REGION Network 3: Release drive
   //
         O     #Temp_IO_Status.Switch_Drive_ON_OFF;
         O     #IN_Request_Filling;
         O     #IN_Request_Feedpump;
         O     #IN_Request_Cooling;
         O     #IN_Request_Heating;
         A     #IN_Release;
         =     #Temp_ReleaseDrive;
END_REGION

REGION Network 4: Faults
         A     #IN_Reset_fault;
         R     #Temp_IO_Fault.FLT_Motorprotection;
         R     #Temp_IO_Fault.FLT_FrequencyConverter;
         R     #Temp_IO_Fault.FLT_MaxP_MaxLTripTray;
         R     #Temp_IO_Fault.FLT_Dryrunsafety;
         R     #Temp_IO_Fault.FLT_wrong_Timevalue;

         A     #IN_Fault_Motorprotection;
         S     #Temp_IO_Fault.FLT_Motorprotection;
         S     #Temp_IO_Status.Reset_Intervall;
   //
         A     #IN_ControlVoltage;
         AN    #Temp_IO_Fault.FLT_wrong_Timevalue;
         AN    #Temp_IO_Status.Start_Startupdelay;
         L     S5T#5S;
         SD    #IN_TimerStartUpFConv;
   //
         A     #IN_TimerStartUpFConv;
         AN    #IN_FaultFreqConverter;
         A     #Temp_ReleaseDrive;
         A     #Temp_IO_Status.Config_bit_with_FC;
         S     #Temp_IO_Fault.FLT_FrequencyConverter;
         S     #Temp_IO_Status.Reset_Intervall;
   //
         AN    #IN_MaxPressure_MaxLTray;
         A     #Temp_ReleaseDrive;
         S     #Temp_IO_Fault.FLT_MaxP_MaxLTripTray;
         S     #Temp_IO_Status.Reset_Intervall;
   //
         AN    #IN_DryRun;
         A     #Temp_ReleaseDrive;
         S     #Temp_IO_Fault.FLT_Dryrunsafety;
         S     #Temp_IO_Status.Reset_Intervall;
END_REGION

REGION Network 5: Time handle
   // Es werden die Absolutwerte der Zeiten berechnet um sie dann vergleichen zu 
   // können. Intervallzeiten sind minimal 10sec. Sonst Störung "Zeitwert falsch"!
   // Bei Spaltfiltern max Laufzeit 20sec.,Min Pausenzeit 300sec.und kein Dauerbetrieb
   // möglich!
         SET;
         R     #Temp_IO_Fault.FLT_wrong_Timevalue;
   //
         L     #IN_DW_RunTime;
         T     #Temp_RunTime;
         L     #IN_DW_PauseTime;
         T     #Temp_PauseTime;
   //
   // Absolutwerte berechnen
   //
         CALL  T_CONV
         ( IN  := #Temp_RunTime,
           OUT := #Temp_Runtime_ms
         );
   //
         CALL  T_CONV
         ( IN  := #Temp_PauseTime,
           OUT := #Temp_Pausetime_ms
         );
   //
         SET;
         R     #Temp_IO_Status.No_Pausetime;
   //
         L     #Temp_Runtime_ms;
         L     0;
         ==I;
         O(;
         L     #Temp_Pausetime_ms;
         L     0;
         ==I;
         );
         AN    #Temp_IO_Status.Config_bit_split;  // Bei Spaltfilter immer mit Intervall
         S     #Temp_IO_Status.No_Pausetime;
   //
   // Zeiten limitieren
   //
         A     #Temp_IO_Status.Config_bit_split;  // Bei Spaltfilter Kontrolle auf spezielle Min und Maxwerte
         JC    nLi2;
   //
         L     #Temp_Runtime_ms;
         L     10000;  // 10 sec
         <D;
         S     #Temp_IO_Fault.FLT_wrong_Timevalue;  // Antrieb STOP!!!
         JCN   nLi1;
         L     S5T#10S;
         T     #Temp_RunTime;
   //
   nLi1: L     #Temp_Pausetime_ms;
         L     10000;  // 10.0 sec
         <D;
         S     #Temp_IO_Fault.FLT_wrong_Timevalue;  // Antrieb STOP!!!
         JCN   nLi3;
         L     S5T#10S;
         T     #Temp_PauseTime;
         JU    nLi3;
   //
   // Sonderteil für Spaltfilter
   nLi2: L     #Temp_Runtime_ms;
         L     20000;  // 20.0 sec
         >D;
         S     #Temp_IO_Fault.FLT_wrong_Timevalue;  // Antrieb STOP!!!
         JCN   KfS1;
         L     S5T#20S;
         T     #Temp_RunTime;
   KfS1: L     #Temp_Pausetime_ms;
         L     L#300000;  // 300.0 sec
         <D;
         S     #Temp_IO_Fault.FLT_wrong_Timevalue;  // Antrieb STOP!!!
         JCN   nLi3;
         L     S5T#5M;
         T     #Temp_PauseTime;
   //
   nLi3: NOP   0;
         A     #Temp_IO_Status.No_Pausetime;  // Wenn eh eine zeit null dann andere egal!
         R     #Temp_IO_Fault.FLT_wrong_Timevalue;
END_REGION

REGION Network 6: Reset Intervall / Angefordert setzen
         O     #Temp_IO_Status.No_Pausetime;
         S     #Temp_IO_Status.Reset_Intervall;
   //
         ON    #Temp_ReleaseDrive;
         ON    #IN_Release;
         O     #Temp_IO_Status.Reset_Intervall;
         R     #Temp_IO_Status.Run;
         R     #Temp_IO_Status.Pause;
         R     #Temp_IO_Status.Reset_Intervall;
END_REGION

REGION Network 7: Wiedereinschaltsperre
         ON    #IN_ControlVoltage;
         FP    #Temp_IO_Status.Ramp_CVoltage_Off;
         S     #Temp_IO_Status.Start_Startupdelay;
         R     #Temp_IO_Status.Disable_Start;
         R     #IN_TimerDrive;
   //
         ON    #Temp_IO_Status.Config_bit_with_FC;
         O     #IN_TimerDrive;
         A     #Temp_IO_Status.Start_Startupdelay;
         R     #Temp_IO_Status.Disable_Start;
         R     #Temp_IO_Status.Start_Startupdelay;
   //
         A     #Temp_IO_Status.Start_Startupdelay;
         JCN   Lauf;
   //
         A     #Temp_IO_Status.Disable_Start;
         L     S5T#10S;
         SD    #IN_TimerDrive;
   //
         SET;
         S     #Temp_IO_Status.Disable_Start;
   //
         A     #IN_TimerDrive;
         A     #Temp_IO_Status.Start_Startupdelay;
         R     #Temp_IO_Status.Start_Startupdelay;
         R     #Temp_IO_Status.Disable_Start;
END_REGION

REGION Network 8: Laufzeit
   Lauf: NOP   0;
         A     #Temp_ReleaseDrive;
         AN    #Temp_IO_Status.Pause;
         AN    #Temp_IO_Status.Start_Startupdelay;
         JCN   Paus;
   //
         A     #Temp_IO_Status.Run;
         L     #Temp_RunTime;
         SD    #IN_TimerDrive;
   //
         SET;
         S     #Temp_IO_Status.Run;
   //
         A     #IN_TimerDrive;
         JCN   Ausg;
         SET;
         R     #Temp_IO_Status.Run;
         R     #IN_TimerDrive;
END_REGION

REGION Network 9: Pause
   Paus: NOP   0;
         A     #Temp_ReleaseDrive;
         AN    #Temp_IO_Status.Run;
         AN    #Temp_IO_Status.Start_Startupdelay;
         JCN   Ausg;
   //
         A     #Temp_IO_Status.Pause;
         L     #Temp_PauseTime;
         SD    #IN_TimerDrive;
   //
         SET;
         S     #Temp_IO_Status.Pause;
   //
         A     #IN_TimerDrive;
         JCN   Ausg;
         SET;
         R     #Temp_IO_Status.Pause;
         R     #IN_TimerDrive;
END_REGION

REGION Network 10: Output mainscontactor
   Ausg: NOP   0;
   //
         A(;
   //
         A     #IN_ControlVoltage;  // generell Eingeschaltet mit FU
         A     #Temp_IO_Status.Config_bit_with_FC;
         AN    #Temp_IO_Status.Start_Startupdelay;
   //
         O(;
         A     #Temp_IO_Status.Run;  // generell Eingeschaltet ohne FU
         O     #Temp_IO_Status.No_Pausetime;
         A     #Temp_IO_Status.Switch_Drive_ON_OFF;
         A(;
         AN    #Temp_IO_Fault.FLT_Dryrunsafety;
         O     #Temp_IO_Status.Config_bit_split;
         );
         AN    #Temp_IO_Status.Config_bit_with_FC;
         );
   //
         O(;
         A     #IN_Request_Filling;  // Befuellen als Füllpumpe
         A     #Temp_IO_Status.Config_bit_char;
         );
   //
         O(;
         O     #Temp_IO_Status.No_Pausetime;  // Befuellen aber normal konfiguriert
         O     #Temp_IO_Status.Run;
         A     #IN_Request_Filling;
         AN    #Temp_IO_Fault.FLT_Dryrunsafety;
         A     #Temp_IO_Status.Config_bit_normal;
         );
   //
         O(;
         A     #IN_Request_Filling;  // aber auch beim Befüllen
         AN    #Temp_IO_Fault.FLT_Dryrunsafety;
         A     #Temp_IO_Status.Run;
         O     #IN_Request_Feedpump;  // Speisen
         A     #Temp_IO_Status.config_bit_feed;
         );
   //
         O(;
         A     #IN_Request_Heating;  // Beim Heizen mit Intervall
         A(;
         O     #Temp_IO_Status.Run;
         O     #Temp_IO_Status.No_Pausetime;
         );
         O     #IN_Request_Cooling;  // Kühlen ohne Intervall, damit WT nicht einfriert
         AN    #Temp_IO_Status.Config_bit_with_FC;
         AN    #Temp_IO_Status.Config_bit_split;
         AN    #Temp_IO_Fault.FLT_Dryrunsafety;
         );
   //
         );
   //
         A(;
         A     #IN_Release;
         AN    #Temp_IO_Fault.FLT_wrong_Timevalue;
         AN    #Temp_IO_Fault.FLT_MaxP_MaxLTripTray;
         O     #Temp_IO_Status.Config_bit_with_FC;  // Wenn FU dann immer an!
         );
         AN    #Temp_IO_Fault.FLT_Motorprotection;
         AN    #Temp_IO_Fault.FLT_Dryrunsafety;
   //
         =     #OUT_MainsContactor;
         =     #Temp_MainsContactor;
END_REGION

REGION Network 11: Ouput release frequency converter
         O     #Temp_IO_Status.No_Pausetime;
         O     #Temp_IO_Status.Run;
         O     #IN_Request_Feedpump;
         A     #IN_Release;
         A     #Temp_MainsContactor;
         A     #Temp_IO_Status.Config_bit_with_FC;
         A(;
         O     #Temp_IO_Status.Switch_Drive_ON_OFF;
         O     #IN_Request_Feedpump;
         );
         AN    #Temp_IO_Fault.FLT_FrequencyConverter;
         A     #IN_FaultFreqConverter;
         =     #OUT_Release_FConverter;
         =     #Temp_Release_FConverter;
END_REGION

REGION Network 12: Error handling
         O     #Temp_IO_Fault.FLT_Motorprotection;
         O     #Temp_IO_Fault.FLT_FrequencyConverter;
         O     #Temp_IO_Fault.FLT_MaxP_MaxLTripTray;
         O     #Temp_IO_Fault.FLT_Dryrunsafety;
         O     #Temp_IO_Fault.FLT_wrong_Timevalue;
         =     #Temp_Fault_Drive;
         =     #Temp_IO_Status.FaultExist;

         O     #Temp_IO_Fault.FLT_Motorprotection;
         O     #Temp_IO_Fault.FLT_FrequencyConverter;
         O     #Temp_IO_Fault.FLT_Dryrunsafety;
         A     #IN_SelectFaultLevel;
         S     #IO_FaultLevel_1;

         O     #Temp_IO_Fault.FLT_Motorprotection;
         O     #Temp_IO_Fault.FLT_FrequencyConverter;
         O     #Temp_IO_Fault.FLT_Dryrunsafety;
         AN    #IN_SelectFaultLevel;
         O;
         O     #Temp_IO_Fault.FLT_MaxP_MaxLTripTray;
         O     #Temp_IO_Fault.FLT_wrong_Timevalue;
         S     #IO_FaultLevel_3;

         O     #Temp_IO_Fault.FLT_Motorprotection;
         FP    #Temp_IO_Status.FLT_Motorprotection;
         S     #IO_NewFault;

         O     #Temp_IO_Fault.FLT_FrequencyConverter;
         FP    #Temp_IO_Status.FLT_FC;
         S     #IO_NewFault;

         O     #Temp_IO_Fault.FLT_MaxP_MaxLTripTray;
         FP    #Temp_IO_Status.FLT_MaxP_MaxLTripTray;
         S     #IO_NewFault;

         O     #Temp_IO_Fault.FLT_Dryrunsafety;
         FP    #Temp_IO_Status.FLT_Dryrunsafety;
         S     #IO_NewFault;

         O     #Temp_IO_Fault.FLT_wrong_Timevalue;
         FP    #Temp_IO_Status.FLT_wrong_Timevalue;
         S     #IO_NewFault;
END_REGION

REGION Network 13: State of drive: 1-> ON; 2->Faulty; 3->Selected but not on
         L     0;
         O     #Temp_Fault_Drive;
         JCN   err;
         L     2;
         JU    tran;
   err:  AN    #Temp_IO_Status.Config_bit_with_FC;
         A     #Temp_MainsContactor;
         O     #Temp_Release_FConverter;
         JCN   anl;
         L     1;
         JU    tran;
   anl:  AN    #Temp_IO_Status.Config_bit_with_FC;
         A     #Temp_MainsContactor;
         O     #Temp_Release_FConverter;
         ON    #Temp_IO_Status.Switch_Drive_ON_OFF;
         JC    tran;
         L     3;
   tran: T     #Temp_IO_Status.State_Drive;
END_REGION

REGION Network 14: Save data
         CALL  BLKMOV
         ( SRCBLK  := #Temp_IO_Status,
           RET_VAL := #ERROR_CODE,
           DSTBLK  := #Anyzeiger1
         );
   //
         CALL  BLKMOV
         ( SRCBLK  := #Temp_IO_Fault,
           RET_VAL := #ERROR_CODE,
           DSTBLK  := #Anyzeiger2
         );
   //
END_REGION
END_FUNCTION

FUNCTION "FC102_Refilling" : Void   // FC102, STL
TITLE = Filling of a tank
{ S7_Optimized_Access := 'FALSE' }
AUTHOR : KT242
FAMILY : RS_KK
NAME : Filling
VERSION : 1.1
// Befüllt wird wahlweise über Niveaugeber "Unten / Oben", "Anzahl Schuesse" oder 
// "Zeit". Das unterschreiten des "IN_Niveau_unten" hat Priorität.
// Vor dem eigentlichen Befüllen läuft die Vorrührzeit ab, sofern sie nicht im 
// Zeit- Zähler- Bedienfeld der Wert "0" eingegeben wurde.
   VAR_INPUT
      IN_Selected : Bool;   // Was this function selected for use?
      IN_ReleaseRefilling : Bool;   // Signal general release refilling
      IN_FillingPumpActive : Bool;   // If filling pump is running filing valve is allowed to open
      IN_WithFillingPump : Bool;   // Select, if filling with filling pump (1) or not (0)
      IN_RecircWeekend : Bool;   // Foaming machine in weekend mode
      IN_FoamingCycleActive : Bool;   // Foaming cycle is active
      IN_PistonActive : Bool;   // Metering unit is a piston
      IN_MH_is_open : Bool;   // Foaming with this component is active // mixinghead open
      IN_ResetFault : Bool;   // Signal quit faults of this funktion block
      IN_MaxLevelTriptray : Bool;   // Max. level of triptray day tank exceeded
      IN_PumpDeselected : Bool;   // Pump(s) of this daytank are deselected -> only fault group 3 on min level
      IN_SetAmountShots : Int;   // Setvalue of shot amout. After this amount of shots refilling starts
      IN_PreAgitatingTime : S5Time;   // Timevalue of pre agitating of a vessel station
      IN_FillingTimeContr : S5Time;   // Timevalue control refilling of daytank
      IN_TimeTillFillingStart : S5Time;   // Timevalue to start refilling after leaving upper level
      IN_Timer_Refilling : Timer;   // Timer of all activities at the function block refilling
   END_VAR
   VAR_OUTPUT
      OUT_V_Preagitating : Bool;   // Output of valve pre agitating of a vessel
      OUT_V_Refilling : Bool;   // Output of valve refilling of tank
      OUT_R_Tankstorage : Bool;   // Output of potential free contakt to an external tank storage
   END_VAR
   VAR_IN_OUT
      IO_Status : ANY;   // State of refilling
      IO_NewFault : Bool;
      IO_FaultLevel_1 : Bool;
      IO_FaultLevel_2 : Bool;
      IO_FaultLevel_3 : Bool;
      IO_Fault : ANY;
   END_VAR
   VAR_TEMP
      Temp_IO_Status : "UDT102_RefillingState";
      ERROR_CODE : Int;   // Error state of systemfunction "BLKMOV" Blockmove
      AnyPointer1 : ANY;   // Pointer to copy thr array "IO_Status" and "Temp_IO_Status"
      AnyPointer2 : ANY;   // Pointer to copy thr array "IO_Status" and "Temp_IO_Status"
      Temp_IO_Fault : "UDT1802_FLT_Tank_Refill";
      Temp_Release : Bool;   // Flag to set release of refilling
      Temp_V_Refilling : Bool;
      Temp_FLTFlag : Bool;
      Temp_FLTstatus : Bool;
   END_VAR
BEGIN

REGION Network 1: Saved data integration
   // nderungen:
   // -------------------------------------------------------------------------------
   // Bei einer Befüllung nach Zeit oder einer Befüllung nach Anzahl Schüssen in kam 
   // es bei Behältern mit nur drei Füllstandsonden (ohne "IN_Niveau_unten") vor das 
   // diese nicht befüllt wurden.
   // Hierbei wurde eine Befüllung nach unterschreiten des Schalters "#IN_Min_Level" 
   // nicht oder verspätet gestartet. 
   // Durch Änderungen im Netzwerk für die normale Befüllung wurde dieses behoben.
   // 
   // Jäger         03.10.2005
   // -------------------------------------------------------------------------------
         LAR1;
         L;
         LAR2;
   //
         L     W[AR2, P#0.0];  // Bytes
         T     W[AR1, P#0.0];
         L     W[AR2, P#2.0];  //Amount of bytes
         T     W[AR1, P#2.0];
         L     W[AR2, P#4.0];  //Block no,
         T     W[AR1, P#4.0];
         L     D[AR2, P#6.0];  //Startadress of datas
         T     D[AR1, P#6.0];
   //
         CALL  BLKMOV
         ( SRCBLK  := #AnyPointer1,
           RET_VAL := #ERROR_CODE,
           DSTBLK  := #Temp_IO_Status
         );
   //
         LAR1;
         L;
         LAR2;
   //
         L     W[AR2, P#0.0];  // Bytes
         T     W[AR1, P#0.0];
         L     W[AR2, P#2.0];  //Amount of bytes
         T     W[AR1, P#2.0];
         L     W[AR2, P#4.0];  //Block no,
         T     W[AR1, P#4.0];
         L     D[AR2, P#6.0];  //Startadress of datas
         T     D[AR1, P#6.0];
   //
         CALL  BLKMOV
         ( SRCBLK  := #AnyPointer2,
           RET_VAL := #ERROR_CODE,
           DSTBLK  := #Temp_IO_Fault
         );
   //
END_REGION

REGION Network 2: Fault handling
         A     #IN_ResetFault;
         ON    #IN_Selected;
         R     #Temp_IO_Fault.FLT_Min_Level;
         R     #Temp_IO_Fault.FLT_Max_Level;
         R     #Temp_IO_Fault.FLT_Fillingtime_to_long;
         R     #Temp_IO_Fault.FLT_Max_Level_Triptray;
         R     #Temp_IO_Fault.FLT_PreWarning_Min_Level;
         R     #Temp_IO_Fault.FLT_Min_Level_Cycle;
         R     #Temp_IO_Fault.FLT_Max_Level_Pistonm;
         R     #Temp_IO_Fault.FLT_Max_Level_Tt_Pistonm;
   //
         ON    #IN_Selected;
         R     #Temp_IO_Status.Fault_Exist;
         R     #Temp_IO_Status.FaultLevel_1;
         R     #Temp_IO_Status.FaultLevel_2;
         R     #Temp_IO_Status.FaultLevel_3;
         JC    Save;
   //
         AN    #Temp_IO_Status.Min_Level;
         AN    #IN_FoamingCycleActive;
         AN    #IN_PumpDeselected;
         AN    #Temp_IO_Fault.FLT_Min_Level;
         S     #Temp_IO_Fault.FLT_Min_Level;
         =     #Temp_FLTFlag;
         A     #Temp_FLTFlag;
         AN    #IN_PumpDeselected;
         S     #IO_FaultLevel_1;
         A     #Temp_FLTFlag;
         A     #IN_PumpDeselected;
         S     #IO_FaultLevel_3;
   //-
         AN    #Temp_IO_Status.Max_Level;
         AN    #IN_PistonActive;
         AN    #Temp_IO_Fault.FLT_Max_Level;
         S     #Temp_IO_Fault.FLT_Max_Level;
         S     #IO_FaultLevel_3;
   //
         AN    #IN_MaxLevelTriptray;
         AN    #IN_PistonActive;
         AN    #Temp_IO_Fault.FLT_Max_Level_Triptray;
         S     #Temp_IO_Fault.FLT_Max_Level_Triptray;
         =     #Temp_FLTFlag;
         A     #Temp_FLTFlag;
         AN    #IN_PumpDeselected;
         S     #IO_FaultLevel_1;
         A     #Temp_FLTFlag;
         A     #IN_PumpDeselected;
         S     #IO_FaultLevel_3;
   //-
         AN    #Temp_IO_Status.Min_Level;
         A     #IN_FoamingCycleActive;
         AN    #IN_PumpDeselected;
         AN    #Temp_IO_Fault.FLT_Min_Level_Cycle;
         S     #Temp_IO_Fault.FLT_Min_Level_Cycle;
         S     #IO_FaultLevel_2;
   //
         AN    #Temp_IO_Status.Max_Level;
         A     #IN_PistonActive;
         AN    #Temp_IO_Fault.FLT_Max_Level_Pistonm;
         S     #Temp_IO_Fault.FLT_Max_Level_Pistonm;
         S     #IO_FaultLevel_1;
   //
         AN    #IN_MaxLevelTriptray;
         A     #IN_PistonActive;
         AN    #Temp_IO_Fault.FLT_Max_Level_Tt_Pistonm;
         S     #Temp_IO_Fault.FLT_Max_Level_Tt_Pistonm;
         S     #IO_FaultLevel_2;
   //-
         A     #Temp_IO_Status.PreWarning_Min_Level;
         AN    #Temp_IO_Fault.FLT_PreWarning_Min_Level;
         S     #Temp_IO_Fault.FLT_PreWarning_Min_Level;
         S     #IO_FaultLevel_3;
   //-
END_REGION

REGION Network 3: Release of refilling
         A     #Temp_IO_Status.Switch_Refilling_ON_OFF;
         A     #IN_ReleaseRefilling;
         AN    #IN_RecircWeekend;
         AN    #Temp_IO_Fault.FLT_Max_Level;
         AN    #Temp_IO_Fault.FLT_Max_Level_Pistonm;
         AN    #Temp_IO_Fault.FLT_Max_Level_Triptray;
         AN    #Temp_IO_Fault.FLT_LevelSensor_broken_wire;
         =     #Temp_Release;
   //
         AN    #Temp_Release;
         R     #Temp_IO_Status.Select_Filling_with_Time;
         R     #IN_Timer_Refilling;
END_REGION

REGION Network 4: Mixinghead is open
         AN    #IN_MH_is_open;  // Start erst nach Schuss
         FP    #Temp_IO_Status.Ramp_MH_open;
         JCN   NSho;
         L     #Temp_IO_Status.Value_No;
         L     1;
         +I;
         T     #Temp_IO_Status.Value_No;
   NSho: NOP   0;
END_REGION

REGION Network 5: Requirement after time
   // Ist eine Zeit >0 vorgegeben wird diese beim Verlassen des Schalters 
   // "IN_Niveau_oben" gestartet.
   // Nach Ablauf der Zeit wird die Befüllung gestartet.
   // Ist kein Schalter "IN_Niveau_unten" vorhanden, muß der Parameter auf true 
   // gesetzt werden.
         ON    #Temp_Release;
         O     #Temp_IO_Status.Select_refilling;
         JC    reg;
   //
         A     #Temp_IO_Status.Select_Filling_with_Time;
         AN    #Temp_IO_Status.Preagitation_runs;
         AN    #Temp_IO_Status.Fillingtime_runs;
         AN    #Temp_IO_Status.Select_refilling;
         L     #IN_TimeTillFillingStart;
         SD    #IN_Timer_Refilling;
   //
         L     #IN_TimeTillFillingStart;  // Zeitwert ausmaskieren
         L     16#0FFF;
         AW;
         L     0;  // Nur wenn Zeit > 0
         >I;
         A     #Temp_IO_Status.Stop_Level_Filling;  // Und oberes Niv verlassen dann aktiviert
         S     #Temp_IO_Status.Select_Filling_with_Time;
   //
         A     #Temp_IO_Status.Select_Filling_with_Time;
         AN    #Temp_IO_Status.Preagitation_runs;
         AN    #Temp_IO_Status.Fillingtime_runs;
         AN    #Temp_IO_Status.Select_refilling;
         A     #IN_Timer_Refilling;
         S     #Temp_IO_Status.Select_refilling;
         R     #IN_Timer_Refilling;
         R     #Temp_IO_Status.Select_Filling_with_Time;
   reg:  NOP   0;
END_REGION

REGION Network 6: Requirement after a amout of shots or by level switch
   // Ist ein Sollwert für Anzahl Schüsse vorgegeben, wird alternativ nach Erreichen 
   // dessen oder bei Unterschreitung des Schalters "IN_Niveau_unten" die Anforderung 
   // gesetzt.
         A(;
         L     #IN_SetAmountShots;  // Sollanzahl > 0
         L     0;
         >I;  //        und
         );
         A(;
         L     #Temp_IO_Status.Value_No;  // Istanzahl >= Sollanzahl
         L     #IN_SetAmountShots;
         >=I;
         );
         ON    #Temp_IO_Status.Start_Level_Filling;
         ON    #Temp_IO_Status.Min_Level;
         AN    #IN_PumpDeselected;
         S     #Temp_IO_Status.Select_refilling;
   //
         ON    #Temp_IO_Status.Stop_Level_Filling;
         JCN   NSta;  // Reguläres Ende
         SET;
         R     #Temp_IO_Status.Select_Filling_with_Time;
         R     #Temp_IO_Status.Select_refilling;
         R     #Temp_IO_Status.Preagitation_runs;
         R     #Temp_IO_Status.Filling_Start;
         R     #Temp_IO_Status.Fillingtime_runs;
         R     #IN_Timer_Refilling;
   //
         L     0;
         T     #Temp_IO_Status.Value_No;
   NSta: NOP   0;
END_REGION

REGION Network 7: Pre stiring of a fessel
         A     #Temp_IO_Status.Select_refilling;
         A     #Temp_Release;
         JCN   Aus;
   //
         A     #Temp_IO_Status.Filling_Start;
         JC    Bef;
   //
         A     #Temp_IO_Status.Preagitation_runs;
         L     #IN_PreAgitatingTime;
         SD    #IN_Timer_Refilling;
   //
         SET;
         S     #Temp_IO_Status.Preagitation_runs;
   //
         A     #IN_Timer_Refilling;
         JCN   Aus;
         SET;
         S     #Temp_IO_Status.Filling_Start;  // Signal an Umwälzpumpe das befüllt werden soll
         R     #IN_Timer_Refilling;
         JU    Aus;
END_REGION

REGION Network 8: Refilling of a Tank
   // Message to PUC if filling is requested but filling pump don't run
   Bef:  A     #Temp_IO_Status.Fillingtime_runs;
         L     #IN_FillingTimeContr;
         SD    #IN_Timer_Refilling;
   //
         A     #IN_FillingPumpActive;  // Erst wenn Pumpe oder Tanklager läuft,
         ON    #IN_WithFillingPump;  // wird tatsächlich befüllt
         A     #Temp_Release;
         S     #Temp_IO_Status.Fillingtime_runs;
   //
         A     #IN_Timer_Refilling;
         JCN   Aus;
         SET;
         AN    #Temp_IO_Fault.FLT_Fillingtime_to_long;
         S     #Temp_IO_Fault.FLT_Fillingtime_to_long;
         S     #IO_FaultLevel_3;
         R     #Temp_IO_Status.Fillingtime_runs;
         R     #Temp_IO_Status.Preagitation_runs;
         R     #IN_Timer_Refilling;
END_REGION

REGION Network 9: Activate the outputs
   Aus:  ON    #Temp_Release;
         ON    #Temp_IO_Status.Select_refilling;
         O     #Temp_IO_Fault.FLT_Fillingtime_to_long;
         R     #Temp_IO_Status.Preagitation_runs;
         R     #Temp_IO_Status.Filling_Start;
         R     #Temp_IO_Status.Fillingtime_runs;
   //
         A     #Temp_IO_Status.Preagitation_runs;
         =     #OUT_V_Preagitating;
   //
         A     #Temp_IO_Status.Filling_Start;
         =     #OUT_R_Tankstorage;  // Es soll befüllt werden auch ans Tanklager
   //
         A     #IN_FillingPumpActive;  // Erst wenn Pumpe oder Tanklager läuft,
         ON    #IN_WithFillingPump;  // wird tatsächlich befüllt
         A     #Temp_IO_Status.Fillingtime_runs;
         =     #OUT_V_Refilling;
         =     #Temp_V_Refilling;
END_REGION

REGION Network 10: Error handling
   //-----
         O     #Temp_IO_Fault.FLT_Max_Level_Triptray;
   //      O     #Temp_IO_Fault.FLT_Min_Level
         O     #Temp_IO_Fault.FLT_Max_Level;
         O     #Temp_IO_Fault.FLT_Max_Level_Pistonm;
         O     #Temp_IO_Fault.FLT_Max_Level_Tt_Pistonm;
         O     #Temp_IO_Fault.FLT_Min_Level_Cycle;
         O     #Temp_IO_Fault.FLT_Fillingtime_to_long;
         O     #Temp_IO_Fault.FLT_LevelSensor_broken_wire;
         O     #Temp_IO_Fault.FLT_PreWarning_Min_Level;
   //-
         O     #Temp_IO_Fault.FLT_NucleationSensor_broken_wire;
         O     #Temp_IO_Fault.FLT_supply_nucleation;
         O     #Temp_IO_Fault.FLT_nucleation;
   //-
         =     #Temp_FLTstatus;

         O     #Temp_FLTstatus;
         O     #Temp_IO_Fault.FLT_Min_Level;
         =     #Temp_IO_Status.Fault_Exist;
   //-----
         O     #Temp_IO_Fault.FLT_Max_Level_Triptray;
         O     #Temp_IO_Fault.FLT_Min_Level;
         AN    #IN_PumpDeselected;
         O     #Temp_IO_Fault.FLT_Max_Level_Pistonm;
         =     #Temp_IO_Status.FaultLevel_1;
         S     #IO_FaultLevel_1;
   //-----
         O     #Temp_IO_Fault.FLT_Max_Level_Tt_Pistonm;
         O     #Temp_IO_Fault.FLT_Min_Level_Cycle;
         =     #Temp_IO_Status.FaultLevel_2;
         S     #IO_FaultLevel_2;
   //-----
         O     #Temp_IO_Fault.FLT_Max_Level_Triptray;
         O     #Temp_IO_Fault.FLT_Min_Level;
         A     #IN_PumpDeselected;
         O     #Temp_IO_Fault.FLT_Fillingtime_to_long;
         O     #Temp_IO_Fault.FLT_Max_Level;
         O     #Temp_IO_Fault.FLT_LevelSensor_broken_wire;
         O     #Temp_IO_Fault.FLT_PreWarning_Min_Level;
         =     #Temp_IO_Status.FaultLevel_3;
         S     #IO_FaultLevel_3;
   //-----
END_REGION

REGION Network 11: State of filling: 1-> ON; 2->Faulty; 3->Selected but not on
         L     0;
         A     #Temp_FLTstatus;
         AN    #Temp_V_Refilling;
         JCN   F_ON;
         L     2;
         JU    tran;
   F_ON: NOP   0;
   //-
         A     #Temp_V_Refilling;
         JCN   anl;
         L     1;
         JU    tran;
   anl:  NOP   0;
   //-
         ON    #Temp_IO_Status.Switch_Refilling_ON_OFF;
         O     #Temp_V_Refilling;
         JC    tran;
         L     3;
   tran: T     #Temp_IO_Status.State_Refilling;
END_REGION

REGION Network 12: Save data
   Save: NOP   0;
         CALL  BLKMOV
         ( SRCBLK  := #Temp_IO_Status,
           RET_VAL := #ERROR_CODE,
           DSTBLK  := #AnyPointer1
         );
   //
         CALL  BLKMOV
         ( SRCBLK  := #Temp_IO_Fault,
           RET_VAL := #ERROR_CODE,
           DSTBLK  := #AnyPointer2
         );
   //
END_REGION
END_FUNCTION

FUNCTION "FC104_FillingSignals" : Void   // FC104, STL
TITLE = Analyses filling leveles and set controlbits of refilling
{ S7_Optimized_Access := 'FALSE' }
NAME : Filling
VERSION : 1.2
// Wertet die Füllstandsanzeige aus, und setzt die bits Niv unten/oben für den 
// Füllbaustein.
   VAR_INPUT
      Tank_exist : Bool;
      Actual_Level_Value : Real;
      IN_With_Level_Probe : Bool;
      IN_With_Triptray : Bool;
      IN_FLT_Level_Probe : Bool;
      IN_Max_Level : Bool;
      IN_Stop_Fill_Level : Bool;
      IN_Start_Fill_Level : Bool;
      IN_Min_Level : Bool;
      IN_Triptray : Bool;
      IN_DrainTank : Bool;
   END_VAR
   VAR_OUTPUT
      OUT_PreWarnMinLevel : Bool;
      OUT_Max_Level : Bool;
      OUT_Stop_Fill_Level : Bool;
      OUT_Start_Fill_Level : Bool;
      OUT_Min_Level : Bool;
      OUT_Enable_Agitator : Bool;
      OUT_Triptray : Bool;
   END_VAR
   VAR_IN_OUT
      IO_TankLevelPar : ANY;
   END_VAR
   VAR_TEMP
      Temp_TankLevelPar : "UDT702_Tank_Level";
      ERROR_CODE : Int;
      Anyzeiger : ANY;   // Pointer to copy thr array "IO_Status" and "Temp_IO_Status"
      Temp_FLT_Level_Probe : Bool;
   END_VAR
BEGIN

REGION Network 1: Saved data integration
   // Änderungen:
   // -------------------------------------------------------------------------------
   // 
   // -------------------------------------------------------------------------------
   //-----
         LAR1;
         L;
         LAR2;
   //-----
         L     16#1002;  // Bytes
         T     W[AR1, P#0.0];
         L     W[AR2, P#2.0];  // Amount of bytes
         T     W[AR1, P#2.0];
         L     W[AR2, P#4.0];  // Block no,
         T     W[AR1, P#4.0];
         L     D[AR2, P#6.0];  // Startadress of datas
         T     D[AR1, P#6.0];
   //-----
         CALL  BLKMOV
         ( SRCBLK  := #Anyzeiger,
           RET_VAL := #ERROR_CODE,
           DSTBLK  := #Temp_TankLevelPar
         );
   //-----
END_REGION

REGION Network 2: detect trip tray
         A     #IN_DrainTank;
         ON    #IN_With_Triptray;
         =     #OUT_Triptray;
END_REGION

REGION Network 3: Check level probe
   //-----
         A     #IN_FLT_Level_Probe;
         A     #IN_With_Level_Probe;
         ON    #Tank_exist;
         R     #OUT_Max_Level;
         R     #OUT_Stop_Fill_Level;
         R     #OUT_Start_Fill_Level;
         R     #OUT_Enable_Agitator;
         R     #OUT_PreWarnMinLevel;
         R     #OUT_Min_Level;
         JC    Out;
   //-----
END_REGION

REGION Network 4: Max Level
   //-----
         ON(;
         L     #Actual_Level_Value;
         L     #Temp_TankLevelPar.Max_Level;
         >R;
         );
         ON    #IN_With_Level_Probe;
         A     #IN_Max_Level;
         =     #OUT_Max_Level;
   //-----
END_REGION

REGION Network 5: Stop filling level
   //-----
         AN(;
         L     #Actual_Level_Value;
         L     #Temp_TankLevelPar.Stop_Level_Filling;
         >R;
         );
         A     #IN_With_Level_Probe;
         O;
         A     #IN_Stop_Fill_Level;
         AN    #IN_With_Level_Probe;
         =     #OUT_Stop_Fill_Level;
   //-----
END_REGION

REGION Network 6: Start filling level
   //-----
         A(;
         L     #Actual_Level_Value;
         L     #Temp_TankLevelPar.Start_Level_Filling;
         >R;
         );
         A     #IN_With_Level_Probe;
         O     #IN_Start_Fill_Level;
         =     #OUT_Start_Fill_Level;
   //-----
END_REGION

REGION Network 7: Enable Agitator level
   //-----
         L     #Temp_TankLevelPar.Stop_Level_Agitator;
         L     #Temp_TankLevelPar.Min_Level;
         >=R;
         JC    LevelAggOK;
         T     #Temp_TankLevelPar.Stop_Level_Agitator;
   LevelAggOK:NOP   0;

         A(;
         L     #Actual_Level_Value;
         L     #Temp_TankLevelPar.Stop_Level_Agitator;
         >=R;
         );
         A     #IN_With_Level_Probe;
         O     #IN_Min_Level;
         =     #OUT_Enable_Agitator;
   //-----
END_REGION

REGION Network 8: Minimum level
   //-----
         A(;
         L     #Actual_Level_Value;
         L     #Temp_TankLevelPar.Min_Level;
         >=R;
         );
         A     #IN_With_Level_Probe;
         O;
         A     #IN_Min_Level;
         O     #IN_DrainTank;
         =     #OUT_Min_Level;
   //-----
END_REGION

REGION Network 9: Warning Minimum level reached
   //-----
         A(;
         L     #Actual_Level_Value;
         L     #Temp_TankLevelPar.Min_Level_Warning;
         <=R;
         );
         A     #IN_With_Level_Probe;
         =     #OUT_PreWarnMinLevel;
   //-----
END_REGION

REGION Network 10: Save data
   //-----
   Out:  NOP   0;
   //-----
         CALL  BLKMOV
         ( SRCBLK  := #Temp_TankLevelPar,
           RET_VAL := #ERROR_CODE,
           DSTBLK  := #Anyzeiger
         );
   //-----
END_REGION
END_FUNCTION

FUNCTION "FC105_Tempering" : Void   // FC105, STL
TITLE = Heating and cooling depending of the mode
{ S7_Optimized_Access := 'FALSE' }
AUTHOR : KT242
NAME : Temp
VERSION : 2.2
   VAR_INPUT
      IN_Exist : Bool;   // Tempering exist
      IN_Release : Bool;   // Release tempering
      IN_Stop_Tempering : Bool;   // Stop tempering if true
      IN_F_Fuse : Bool;   // Fault fuse
      IN_F_Limit : Bool;   // Fault hardware limit reached
      IN_FLT_Ackn : Bool;   // Fault acknowledge
      IN_CoolingRequested : Bool;   // Cooling requested
      IN_HeatingRequested : Bool;   // Heating requested
      IN_actual_Temp : Real;
      IN_set_Temp : Real;
   END_VAR
   VAR_OUTPUT
      Out_act_cooling : Bool;   // Relais heating or cooling
      Out_act_request_cooling : Bool;   // Request of actuator
      Out_act_heating : Bool;   // Relais heating or cooling
      Out_act_request_heating : Bool;   // Request of actuator
   END_VAR
   VAR_IN_OUT
      IO_StateCtrl1 : ANY;   // Controller State of Controller 1
      IO_ValueCtrl1 : ANY;   // Values of Controller 1
      IO_FaultsCtrl1 : ANY;   // Fault bits of Controller 1
      IO_NewFault : Bool;
      IO_FaultLevel_3 : Bool;
   END_VAR
   VAR_TEMP
      Anyzeiger1 : ANY;   // Pointer to copy thr array "IO_Values" and "Temp_IO_Values"
      Anyzeiger2 : ANY;   // Pointer to copy thr array "IO_Status" and "Temp_IO_Status"
      Anyzeiger3 : ANY;
      Temp_IO_Values : "UDT703_TemperingControl";
      Temp_IO_State : "UDT105_Controller_State";
      TEMP_IO_Faults : "UDT1804_FLT_Controller";
      ERROR_CODE : Int;   // Error state of systemfunction "BLKMOV" Blockmove
      Temp_No_Valid_HeatValue : Bool;
      Temp_No_Valid_CoolValue : Bool;
      Temp_No_Settings_Requested : Bool;
      Temp_Cooling_On : Real;
      Temp_Heating_On : Real;
      Temp_Cooling_Off : Real;
      Temp_Heating_Off : Real;
      Temp_Anf_1 : Byte;
      Temp_Anf_2 : Word;
      Temp_Anf_DW : Word;
      Temp_Anf_1_R : Byte;
      Temp_Anf_2_R : Word;
   END_VAR
BEGIN

REGION Network 1: Relais heating or cooling
         A     #IN_Exist;
         JC    strt;
         R     #Out_act_cooling;
         R     #Out_act_request_cooling;
         R     #Out_act_heating;
         R     #Out_act_request_heating;
         R     #Temp_IO_State.Fault_Exist;
         R     #TEMP_IO_Faults.HW_Limit;
         R     #TEMP_IO_Faults.Fuse_TemperingOverLoad;
         R     #TEMP_IO_Faults.lower_limit;
         R     #TEMP_IO_Faults.upper_limit;
         R     #TEMP_IO_Faults.NoSetValue;
         BEU;
   strt: NOP   0;
END_REGION

REGION Network 2: Read Values of Heating and Cooling fromdata block
   //------------------------------------------------------------
   // Copy dataset of controller parameters connected with PV
   //------------------------------------------------------------
         L;
         LAR1;
   // create any pointer of sourcedata block of selected controller
         LAR2;
   //
   // Type of data to be transmitted
         L     W[AR1, P#0.0];  // Datentyp 10 - S7; 02 - Byte
         T     W[AR2, P#0.0];
   // Amount of datas (length od data set)
         L     W[AR1, P#2.0];  // Wiederholfaktor
         T     W[AR2, P#2.0];
   // DB-number
         L     W[AR1, P#4.0];
         T     W[AR2, P#4.0];

         L     16#84;  //LB [AR1,P#6.0]              // Speicherbereich 84 - DB
         T     LB[AR2, P#6.0];

         L     B[AR1, P#7.0];  // Byte Adresse zusammensetzen
         SLW   13;
         T     #Temp_Anf_1;

         L     W[AR1, P#8.0];
         SRW   3;
         L     #Temp_Anf_1;
         OW;
         T     #Temp_Anf_2;

   // Adresspointer; No of dataset controller data
   //      L W [ AR1 , P#2.0 ]        // length in byte
         L     #Temp_Anf_2;
   //      +D
         T     #Temp_Anf_DW;

         L     #Temp_Anf_DW;
         SRW   13;
         T     #Temp_Anf_1_R;  // Berechnung Anfangsbyte

         L     #Temp_Anf_DW;
         SLW   3;
         T     #Temp_Anf_2_R;

   // Adresspointer; dataset of the controller needs to be included
         L     #Temp_Anf_1_R;
         T     LB[AR2, P#7.0];
         L     #Temp_Anf_2_R;
         T     LW[AR2, P#8.0];
   //
         CALL  BLKMOV
         ( SRCBLK  := #Anyzeiger1,
           RET_VAL := #ERROR_CODE,
           DSTBLK  := #Temp_IO_Values
         );

   //------------------------------------------------------------
   // Copy dataset state of controller connected with PV
   //------------------------------------------------------------
         L;
         LAR1;

         LAR2;

   // Type of data to be transmitted
         L     W[AR1, P#0.0];  // Datentyp 10 - S7; 02 - Byte
         T     W[AR2, P#0.0];
   // Amount of datas (length od data set)
         L     W[AR1, P#2.0];  // Wiederholfaktor
         T     W[AR2, P#2.0];
   // DB-number
         L     W[AR1, P#4.0];
         T     W[AR2, P#4.0];

         L     16#84;  // L     LB [AR1,P#6.0]              // Speicherbereich 84 - DB
         T     LB[AR2, P#6.0];

         L     B[AR1, P#7.0];  //Start Adresse des Datenbereichs zusammensetzen
         SLW   13;
         T     #Temp_Anf_1;

         L     W[AR1, P#8.0];
         SRW   3;
         L     #Temp_Anf_1;
         OW;
         T     #Temp_Anf_2;  //Start Adresse des Datenbereichs

   // Adresspointer; No of dataset controller data
   //      L W [ AR1 , P#2.0 ]        // length in byte
         L     #Temp_Anf_2;
   //      +D
         T     #Temp_Anf_DW;

         L     #Temp_Anf_DW;
         SRW   13;
         T     #Temp_Anf_1_R;  // Calculate start byte

         L     #Temp_Anf_DW;
         SLW   3;
         T     #Temp_Anf_2_R;

   // Adresspointer; dataset of the controller needs to be included
         L     #Temp_Anf_1_R;
         T     LB[AR2, P#7.0];
         L     #Temp_Anf_2_R;
         T     LW[AR2, P#8.0];

   //
         CALL  BLKMOV
         ( SRCBLK  := #Anyzeiger2,
           RET_VAL := #ERROR_CODE,
           DSTBLK  := #Temp_IO_State
         );
END_REGION

REGION Network 3: Read state controller faults
   //------------------------------------------------------------
   // Copy dataset faults of controller connected with PV
   //------------------------------------------------------------
         L;
         LAR1;

         LAR2;

   // Type of data to be transmitted
         L     W[AR1, P#0.0];  // Datentyp 10 - S7; 02 - Byte
         T     W[AR2, P#0.0];
   // Amount of datas (length od data set)
         L     W[AR1, P#2.0];  // Wiederholfaktor
         T     W[AR2, P#2.0];
   // DB-number
         L     W[AR1, P#4.0];
         T     W[AR2, P#4.0];

         L     16#84;  // L     LB [AR1,P#6.0]              // Speicherbereich 84 - DB
         T     LB[AR2, P#6.0];

         L     B[AR1, P#7.0];  //Start Adresse des Datenbereichs zusammensetzen
         SLW   13;
         T     #Temp_Anf_1;

         L     W[AR1, P#8.0];
         SRW   3;
         L     #Temp_Anf_1;
         OW;
         T     #Temp_Anf_2;  //Start Adresse des Datenbereichs

   // Adresspointer; No of dataset controller data
   //      L W [ AR1 , P#2.0 ]        // length in byte
         L     #Temp_Anf_2;
   //      +D
         T     #Temp_Anf_DW;

         L     #Temp_Anf_DW;
         SRW   13;
         T     #Temp_Anf_1_R;  // Calculate start byte

         L     #Temp_Anf_DW;
         SLW   3;
         T     #Temp_Anf_2_R;

   // Adresspointer; dataset of the controller needs to be included
         L     #Temp_Anf_1_R;
         T     LB[AR2, P#7.0];
         L     #Temp_Anf_2_R;
         T     LW[AR2, P#8.0];

   //
         CALL  BLKMOV
         ( SRCBLK  := #Anyzeiger3,
           RET_VAL := #ERROR_CODE,
           DSTBLK  := #TEMP_IO_Faults
         );
END_REGION

REGION Network 4: Error handling
         A     #IN_FLT_Ackn;
         R     #TEMP_IO_Faults.HW_Limit;
         R     #TEMP_IO_Faults.Fuse_TemperingOverLoad;
         R     #TEMP_IO_Faults.lower_limit;
         R     #TEMP_IO_Faults.upper_limit;
         R     #TEMP_IO_Faults.NoSetValue;

   // Sets fault if min.temp > 0 and act.temp < min.temp
         A(;
         L     #Temp_IO_Values.Min_Temp;
         L     0.0;
         >R;
         );
         A(;
         L     #IN_actual_Temp;
         L     #Temp_IO_Values.Min_Temp;
         <R;
         );
         A     #Temp_IO_State.Switch_Temp_ON_OFF;
         AN    #TEMP_IO_Faults.lower_limit;
         S     #IO_NewFault;
         S     #TEMP_IO_Faults.lower_limit;

   // Sets fault if man.temp > 0 and act.temp > max.temp
         A(;
         L     #Temp_IO_Values.Max_Temp;
         L     0.0;
         >R;
         );
         A(;
         L     #IN_actual_Temp;
         L     #Temp_IO_Values.Max_Temp;
         >R;
         );
         A     #Temp_IO_State.Switch_Temp_ON_OFF;
         AN    #TEMP_IO_Faults.upper_limit;
         S     #IO_NewFault;
         S     #TEMP_IO_Faults.upper_limit;

         AN    #IN_F_Fuse;
         A     #IN_HeatingRequested;
         A     #Temp_IO_State.Switch_Temp_ON_OFF;
         AN    #TEMP_IO_Faults.Fuse_TemperingOverLoad;
         S     #IO_NewFault;
         S     #TEMP_IO_Faults.Fuse_TemperingOverLoad;

         A     #IN_F_Limit;
         A     #Temp_IO_State.Switch_Temp_ON_OFF;
         AN    #TEMP_IO_Faults.HW_Limit;
         S     #IO_NewFault;
         S     #TEMP_IO_Faults.HW_Limit;

         A(;
         L     #IN_set_Temp;
         L     0.0;
         ==D;
         );
         A     #Temp_IO_State.Switch_Temp_ON_OFF;
         AN    #TEMP_IO_Faults.NoSetValue;
         S     #IO_NewFault;
         S     #TEMP_IO_Faults.NoSetValue;

         O     #TEMP_IO_Faults.HW_Limit;
         O     #TEMP_IO_Faults.Fuse_TemperingOverLoad;
         O     #TEMP_IO_Faults.lower_limit;
         O     #TEMP_IO_Faults.upper_limit;
         O     #TEMP_IO_Faults.NoSetValue;
         S     #IO_FaultLevel_3;
END_REGION

REGION Network 5: Select all fault messages of the temperatur controler
   //-----
         O     #TEMP_IO_Faults.Sensor_FLT_broken_wire;
         O     #TEMP_IO_Faults.Warning_limit_plus;
         O     #TEMP_IO_Faults.Warning_limit_minus;
         O     #TEMP_IO_Faults.Alarm_limit_plus;
         O     #TEMP_IO_Faults.Alarm_limit_minus;
         O     #TEMP_IO_Faults.Controller_at_limit;
   //-
         O     #TEMP_IO_Faults.HW_Limit;
         O     #TEMP_IO_Faults.Fuse_TemperingOverLoad;
         O     #TEMP_IO_Faults.lower_limit;
         O     #TEMP_IO_Faults.upper_limit;
         O     #TEMP_IO_Faults.NoSetValue;
   //-
         O     #TEMP_IO_Faults.Fuse_TemperingUnit;
   //-
         =     #Temp_IO_State.Fault_Exist;
   //-----
END_REGION

REGION Network 6: Test the values
         O(;
         L     #Temp_IO_Values.Dif_Cooling_ON;
         L     0.0;
         ==R;
         );
         O(;
         L     #Temp_IO_Values.Dif_Cooling_ON;
         L     #Temp_IO_Values.Dif_Cooling_OFF;
         <R;
         );
         =     #Temp_No_Valid_CoolValue;

         O(;
         L     #Temp_IO_Values.Dif_Heating_ON;
         L     0.0;
         ==R;
         );
         O(;
         L     #Temp_IO_Values.Dif_Heating_ON;
         L     #Temp_IO_Values.Dif_Heating_OFF;
         <R;
         );
         =     #Temp_No_Valid_HeatValue;
END_REGION

REGION Network 7: Calculate limits

         L     #IN_set_Temp;
         L     #Temp_IO_Values.Dif_Heating_ON;
         -R;
         T     #Temp_Heating_On;

         L     #IN_set_Temp;
         L     #Temp_IO_Values.Dif_Heating_OFF;
         -R;
         T     #Temp_Heating_Off;

         L     #IN_set_Temp;
         L     #Temp_IO_Values.Dif_Cooling_ON;
         +R;
         T     #Temp_Cooling_On;

         L     #IN_set_Temp;
         L     #Temp_IO_Values.Dif_Cooling_OFF;
         +R;
         T     #Temp_Cooling_Off;
END_REGION

REGION Network 8: Cooling mode
         AN    #IN_CoolingRequested;
         O     #TEMP_IO_Faults.NoSetValue;
         R     #Temp_IO_State.CoolingRequest;
         JC    OUTC;

         L     #IN_actual_Temp;  // Actual Value > Switch ON value
         L     #Temp_Cooling_On;
         >R;
         S     #Temp_IO_State.CoolingRequest;

         O(;
         L     #IN_actual_Temp;
         L     #Temp_Cooling_Off;
         <=R;
         );
         O(;
         L     #IN_actual_Temp;
         L     #Temp_IO_Values.Min_Temp;
         <R;
         );
         O     #Temp_No_Valid_CoolValue;
         ON    #Temp_IO_State.Switch_Temp_ON_OFF;
         R     #Temp_IO_State.CoolingRequest;

   OUTC: A     #Temp_IO_State.CoolingRequest;
         =     #Out_act_request_cooling;

         A     #IN_Release;
         AN    #IN_Stop_Tempering;
         A     #Temp_IO_State.CoolingRequest;
         AN    #TEMP_IO_Faults.lower_limit;
         =     #Out_act_cooling;
         =     #Temp_IO_State.CoolingActive;
END_REGION

REGION Network 9: Heating mode
   // Kühlen ist dominant
         AN    #IN_HeatingRequested;
         O     #TEMP_IO_Faults.NoSetValue;
         R     #Temp_IO_State.HeatingRequest;
         JC    OUTH;

         L     #IN_actual_Temp;  // Actual Temp < Switch ON value
         L     #Temp_Heating_On;
         <R;
         S     #Temp_IO_State.HeatingRequest;

         A(;
         L     #IN_actual_Temp;
         L     #Temp_IO_Values.Max_Temp;
         >R;
         );
         A(;
         L     #Temp_IO_Values.Max_Temp;
         L     0.0;
         >R;
         );
         O(;
         L     #IN_actual_Temp;
         L     #Temp_Heating_Off;
         >=R;
         );
         O     #Temp_No_Valid_HeatValue;
         O     #Temp_IO_State.CoolingRequest;
         ON    #Temp_IO_State.Switch_Temp_ON_OFF;
         R     #Temp_IO_State.HeatingRequest;

   OUTH: A     #Temp_IO_State.HeatingRequest;
         =     #Out_act_request_heating;

         A     #IN_Release;
         AN    #IN_Stop_Tempering;
         A     #Temp_IO_State.HeatingRequest;
         AN    #TEMP_IO_Faults.Fuse_TemperingOverLoad;
         AN    #TEMP_IO_Faults.HW_Limit;
         AN    #TEMP_IO_Faults.upper_limit;
         =     #Out_act_heating;
         =     #Temp_IO_State.HeatingActive;
END_REGION

REGION Network 10: State tempering 1: ON; 2:error; 3:Selected but not ON
         L     0;
         O     #TEMP_IO_Faults.Fuse_TemperingOverLoad;
         O     #TEMP_IO_Faults.HW_Limit;
         JCN   F_ON;
         L     2;
         JU    tran;
   F_ON: O     #Temp_IO_State.HeatingActive;
         O     #Temp_IO_State.CoolingActive;
         JCN   anl;
         L     1;
         JU    tran;
   anl:  ON    #Temp_IO_State.Switch_Temp_ON_OFF;
         O     #Temp_IO_State.HeatingActive;
         O     #Temp_IO_State.CoolingActive;
         JC    tran;
         L     3;
   tran: T     #Temp_IO_State.State_Temp;
END_REGION

REGION Network 11: Save Values
         CALL  BLKMOV
         ( SRCBLK  := #Temp_IO_State,
           RET_VAL := #ERROR_CODE,
           DSTBLK  := #Anyzeiger2
         );

         CALL  BLKMOV
         ( SRCBLK  := #TEMP_IO_Faults,
           RET_VAL := #ERROR_CODE,
           DSTBLK  := #Anyzeiger3
         );
END_REGION
END_FUNCTION

FUNCTION "FC106_Vacuum" : Void   // FC106, STL
TITLE = Vacuum pump of day tank
{ S7_Optimized_Access := 'FALSE' }
AUTHOR : KT242
NAME : Vakuum
VERSION : 1.0
// Bei Vorwahl "mit Vakuum" und der Druckschalter meldet "Vakuum nicht erreicht" 
// wird zuerst die Vakuumpumpe angesteuert und 0,5sec. später das Absperrventil.
// Meldet der Druckschalter "Vakuum erreicht", dann wird zuerst das Absperrventil 
// abgesteuert und 0,5sec. später die Vakuumpumpe.
// Bei Vorwahl "mit Vordruck" oder keine gültige Betriebsart erfolgt keine 
// Ansteuerung der Ventile.
   VAR_INPUT
      IN_Release : Bool;   // General release of vacuum function
      IN_P_Vacuum : Bool;   // Input of vacuum pressure switch
      IN_Timer_delay_Lock : Timer;   // Timer delay of locking valve
      IN_Timer_delay_Pumpe : Timer;   // Timer delay switch of vacuum pump after vacuum pressure reached
   END_VAR
   VAR_OUTPUT
      OUT_V_Lock_Vacuum : Bool;   // Output locking valve vacuums
      OUT_V_Pump_Vacuum : Bool;   // Output vakuum pump
      OUT_H_Vacuum_active : Bool;   // Indicator vakuum pump active
   END_VAR
   VAR_IN_OUT
      IO_Status : "UDT106_Vacuum_Status";
   END_VAR
BEGIN

REGION Network 1: Select without vacuum -> with pre pressure
         ON    #IO_Status.Switch_Vacuum_ON_OFF;
         ON    #IN_Release;
         JCN   VAK;
   //
         R     #OUT_V_Lock_Vacuum;
         R     #OUT_V_Pump_Vacuum;
         R     #OUT_H_Vacuum_active;
   //
         CLR;
         L     0;
         SD    #IN_Timer_delay_Lock;
         SD    #IN_Timer_delay_Pumpe;

         ON    #IO_Status.Switch_Vacuum_ON_OFF;
         JC    NoAktivStat;
         L     3;
   NoAktivStat:NOP   0;
         T     #IO_Status.Status_Vacuum;
         BEU;
END_REGION
